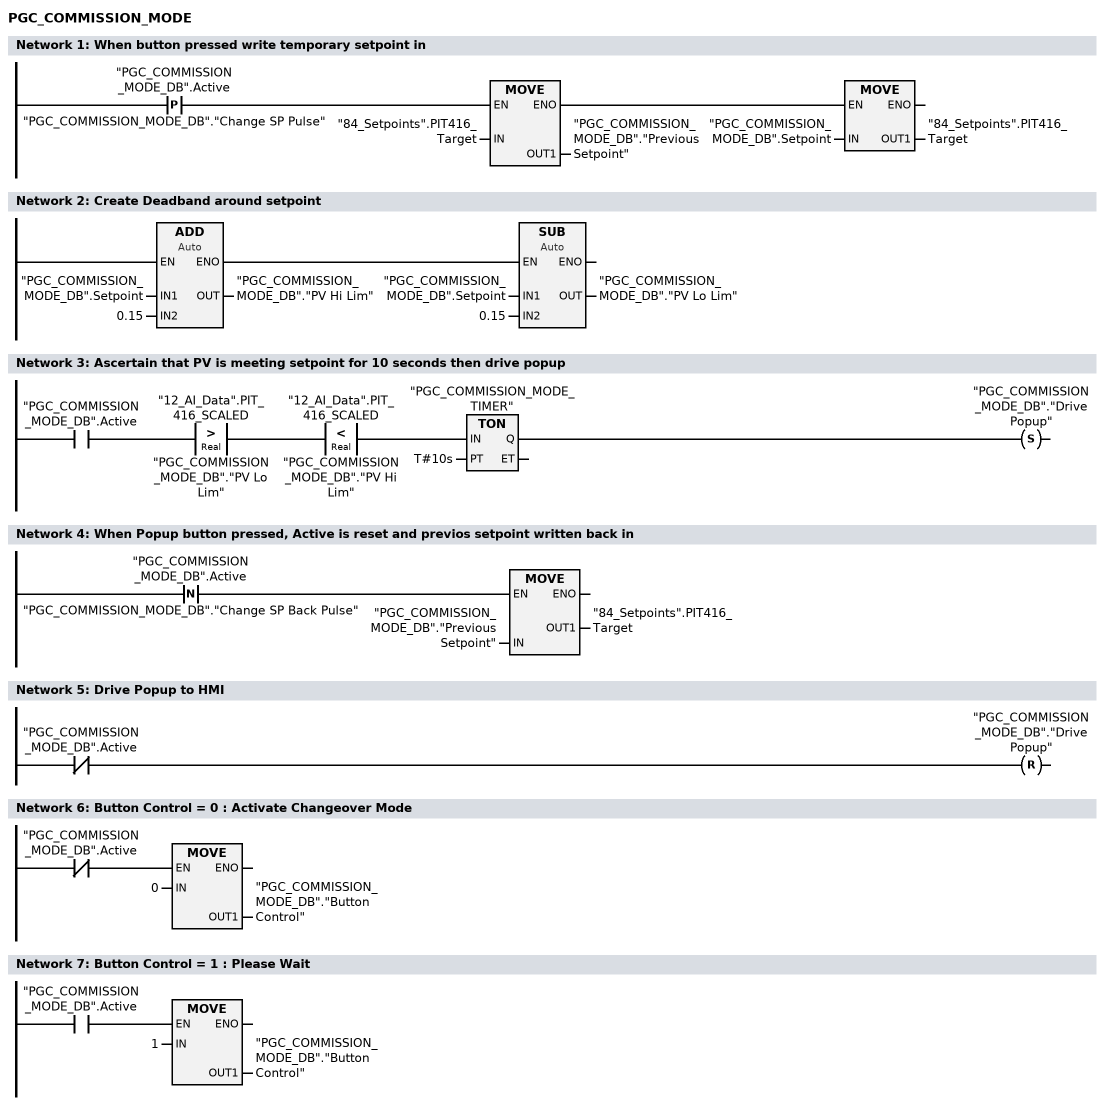
   RUNG wire#powerrail
      P_Contact(operand := "PGC_COMMISSION_MODE_DB".Active, bit := "PGC_COMMISSION_MODE_DB"."Change SP Pulse")
      Move(in := "84_Setpoints".PIT416_Target, out1 => "PGC_COMMISSION_MODE_DB"."Previous Setpoint")
      Move(in := "PGC_COMMISSION_MODE_DB".Setpoint, out1 => "84_Setpoints".PIT416_Target)
   END_RUNG
   // the same network as SCL:
   #_w1 := "PGC_COMMISSION_MODE_DB".Active AND NOT "PGC_COMMISSION_MODE_DB"."Change SP Pulse";   // rising edge of "PGC_COMMISSION_MODE_DB".Active
   "PGC_COMMISSION_MODE_DB"."Change SP Pulse" := "PGC_COMMISSION_MODE_DB".Active;
   IF #_w1 THEN
       "PGC_COMMISSION_MODE_DB"."Previous Setpoint" := "84_Setpoints".PIT416_Target;
       "84_Setpoints".PIT416_Target := "PGC_COMMISSION_MODE_DB".Setpoint;
   END_IF;
END_REGION

REGION Network 2: Create Deadband around setpoint
   RUNG wire#powerrail
      Add(in1 := "PGC_COMMISSION_MODE_DB".Setpoint, in2 := 0.15, out => "PGC_COMMISSION_MODE_DB"."PV Hi Lim")
      Sub(in1 := "PGC_COMMISSION_MODE_DB".Setpoint, in2 := 0.15, out => "PGC_COMMISSION_MODE_DB"."PV Lo Lim")
   END_RUNG
   // the same network as SCL:
   "PGC_COMMISSION_MODE_DB"."PV Hi Lim" := "PGC_COMMISSION_MODE_DB".Setpoint + 0.15;
   "PGC_COMMISSION_MODE_DB"."PV Lo Lim" := "PGC_COMMISSION_MODE_DB".Setpoint - 0.15;
END_REGION

REGION Network 3: Ascertain that PV is meeting setpoint for 10 seconds then drive popup
   "PGC_COMMISSION_MODE_TIMER".TON(IN := "PGC_COMMISSION_MODE_DB".Active AND ("12_AI_Data".PIT_416_SCALED > "PGC_COMMISSION_MODE_DB"."PV Lo Lim") AND ("12_AI_Data".PIT_416_SCALED < "PGC_COMMISSION_MODE_DB"."PV Hi Lim"),
                           PT := T#10s);
   IF "PGC_COMMISSION_MODE_TIMER".Q THEN "PGC_COMMISSION_MODE_DB"."Drive Popup" := TRUE; END_IF;
END_REGION

REGION Network 4: When Popup button pressed, Active is reset and previos setpoint written back in
   RUNG wire#powerrail
      N_Contact(operand := "PGC_COMMISSION_MODE_DB".Active, bit := "PGC_COMMISSION_MODE_DB"."Change SP Back Pulse")
      Move(in := "PGC_COMMISSION_MODE_DB"."Previous Setpoint", out1 => "84_Setpoints".PIT416_Target)
   END_RUNG
   // the same network as SCL:
   #_w1 := NOT "PGC_COMMISSION_MODE_DB".Active AND "PGC_COMMISSION_MODE_DB"."Change SP Back Pulse";   // falling edge of "PGC_COMMISSION_MODE_DB".Active
   "PGC_COMMISSION_MODE_DB"."Change SP Back Pulse" := "PGC_COMMISSION_MODE_DB".Active;
   IF #_w1 THEN "84_Setpoints".PIT416_Target := "PGC_COMMISSION_MODE_DB"."Previous Setpoint"; END_IF;
END_REGION

REGION Network 5: Drive Popup to HMI
   RUNG wire#powerrail
      I_Contact( "PGC_COMMISSION_MODE_DB".Active )
      R_Coil( "PGC_COMMISSION_MODE_DB"."Drive Popup" )
   END_RUNG
   // the same network as SCL:
   IF NOT "PGC_COMMISSION_MODE_DB".Active THEN "PGC_COMMISSION_MODE_DB"."Drive Popup" := FALSE; END_IF;
END_REGION

REGION Network 6: Button Control = 0 : Activate Changeover Mode
   RUNG wire#powerrail
      I_Contact( "PGC_COMMISSION_MODE_DB".Active )
      Move(in := 0, out1 => "PGC_COMMISSION_MODE_DB"."Button Control")
   END_RUNG
   // the same network as SCL:
   IF NOT "PGC_COMMISSION_MODE_DB".Active THEN "PGC_COMMISSION_MODE_DB"."Button Control" := 0; END_IF;
END_REGION

REGION Network 7: Button Control = 1 : Please Wait
   RUNG wire#powerrail
      Contact( "PGC_COMMISSION_MODE_DB".Active )
      Move(in := 1, out1 => "PGC_COMMISSION_MODE_DB"."Button Control")
   END_RUNG
   // the same network as SCL:
   IF "PGC_COMMISSION_MODE_DB".Active THEN "PGC_COMMISSION_MODE_DB"."Button Control" := 1; END_IF;
END_REGION
END_FUNCTION

// folder: 90 - 99 Manual Functions

FUNCTION "90_Manual_Control" : Void   // FC90, LAD
TITLE = Manual Control
{ S7_Optimized_Access := 'TRUE' }
AUTHOR : JHT
VERSION : 0.1
// Code for manual operation of equipment
   VAR_TEMP   // added for the SCL form of the ladder/FBD networks
      _w1 : Bool;
      _w2 : Bool;
      _w3 : Bool;
      _w4 : Bool;
      _w5 : Bool;
      _w6 : Bool;
   END_VAR
BEGIN

REGION Network 1: Q136.0 - Fresh Water Fill Valve Control (CV358)
   // True = Activate, False = NOT
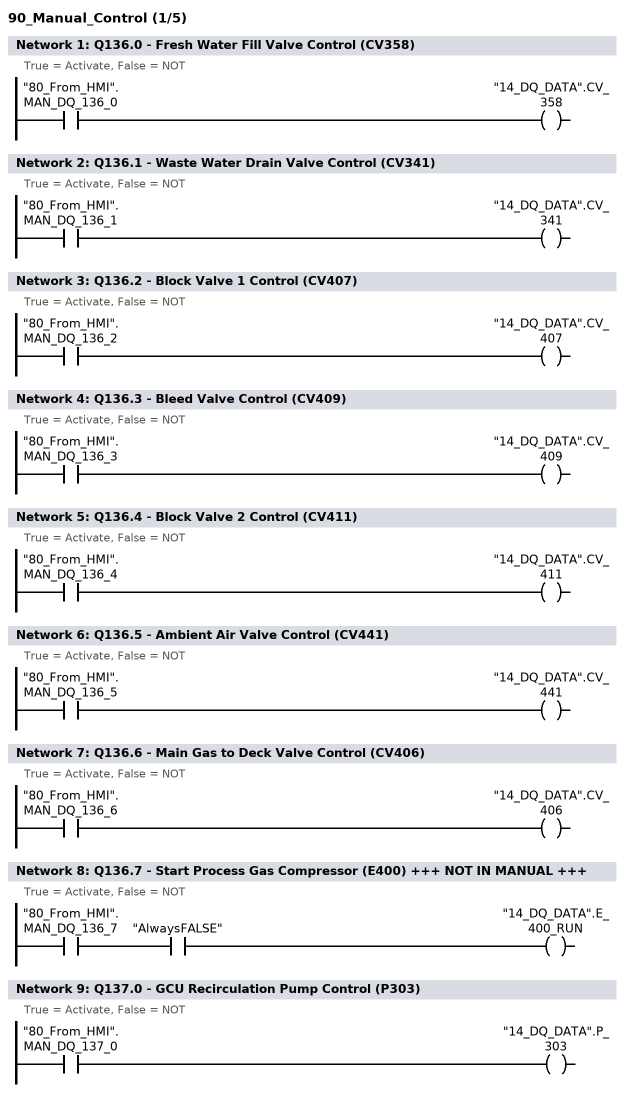
   RUNG wire#powerrail
      Contact( "80_From_HMI".MAN_DQ_136_0 )
      Coil( "14_DQ_DATA".CV_358 )
   END_RUNG
   // the same network as SCL:
   "14_DQ_DATA".CV_358 := "80_From_HMI".MAN_DQ_136_0;
END_REGION

REGION Network 2: Q136.1 - Waste Water Drain Valve Control (CV341)
   // True = Activate, False = NOT
   RUNG wire#powerrail
      Contact( "80_From_HMI".MAN_DQ_136_1 )
      Coil( "14_DQ_DATA".CV_341 )
   END_RUNG
   // the same network as SCL:
   "14_DQ_DATA".CV_341 := "80_From_HMI".MAN_DQ_136_1;
END_REGION

REGION Network 3: Q136.2 - Block Valve 1 Control (CV407)
   // True = Activate, False = NOT
   RUNG wire#powerrail
      Contact( "80_From_HMI".MAN_DQ_136_2 )
      Coil( "14_DQ_DATA".CV_407 )
   END_RUNG
   // the same network as SCL:
   "14_DQ_DATA".CV_407 := "80_From_HMI".MAN_DQ_136_2;
END_REGION

REGION Network 4: Q136.3 - Bleed Valve Control (CV409)
   // True = Activate, False = NOT
   RUNG wire#powerrail
      Contact( "80_From_HMI".MAN_DQ_136_3 )
      Coil( "14_DQ_DATA".CV_409 )
   END_RUNG
   // the same network as SCL:
   "14_DQ_DATA".CV_409 := "80_From_HMI".MAN_DQ_136_3;
END_REGION

REGION Network 5: Q136.4 - Block Valve 2 Control (CV411)
   // True = Activate, False = NOT
   RUNG wire#powerrail
      Contact( "80_From_HMI".MAN_DQ_136_4 )
      Coil( "14_DQ_DATA".CV_411 )
   END_RUNG
   // the same network as SCL:
   "14_DQ_DATA".CV_411 := "80_From_HMI".MAN_DQ_136_4;
END_REGION

REGION Network 6: Q136.5 - Ambient Air Valve Control (CV441)
   // True = Activate, False = NOT
   RUNG wire#powerrail
      Contact( "80_From_HMI".MAN_DQ_136_5 )
      Coil( "14_DQ_DATA".CV_441 )
   END_RUNG
   // the same network as SCL:
   "14_DQ_DATA".CV_441 := "80_From_HMI".MAN_DQ_136_5;
END_REGION

REGION Network 7: Q136.6 - Main Gas to Deck Valve Control (CV406)
   // True = Activate, False = NOT
   RUNG wire#powerrail
      Contact( "80_From_HMI".MAN_DQ_136_6 )
      Coil( "14_DQ_DATA".CV_406 )
   END_RUNG
   // the same network as SCL:
   "14_DQ_DATA".CV_406 := "80_From_HMI".MAN_DQ_136_6;
END_REGION

REGION Network 8: Q136.7 - Start Process Gas Compressor (E400) +++ NOT IN MANUAL +++
   // True = Activate, False = NOT
   RUNG wire#powerrail
      Contact( "80_From_HMI".MAN_DQ_136_7 )
      Contact( "AlwaysFALSE" )
      Coil( "14_DQ_DATA".E_400_RUN )
   END_RUNG
   // the same network as SCL:
   "14_DQ_DATA".E_400_RUN := "80_From_HMI".MAN_DQ_136_7 AND "AlwaysFALSE";
END_REGION

REGION Network 9: Q137.0 - GCU Recirculation Pump Control (P303)
   // True = Activate, False = NOT
   RUNG wire#powerrail
      Contact( "80_From_HMI".MAN_DQ_137_0 )
      Coil( "14_DQ_DATA".P_303 )
   END_RUNG
   // the same network as SCL:
   "14_DQ_DATA".P_303 := "80_From_HMI".MAN_DQ_137_0;
END_REGION

REGION Network 10: Q137.1 - GCU Booster Pump Control (P304)
   // True = Activate, False = NOT
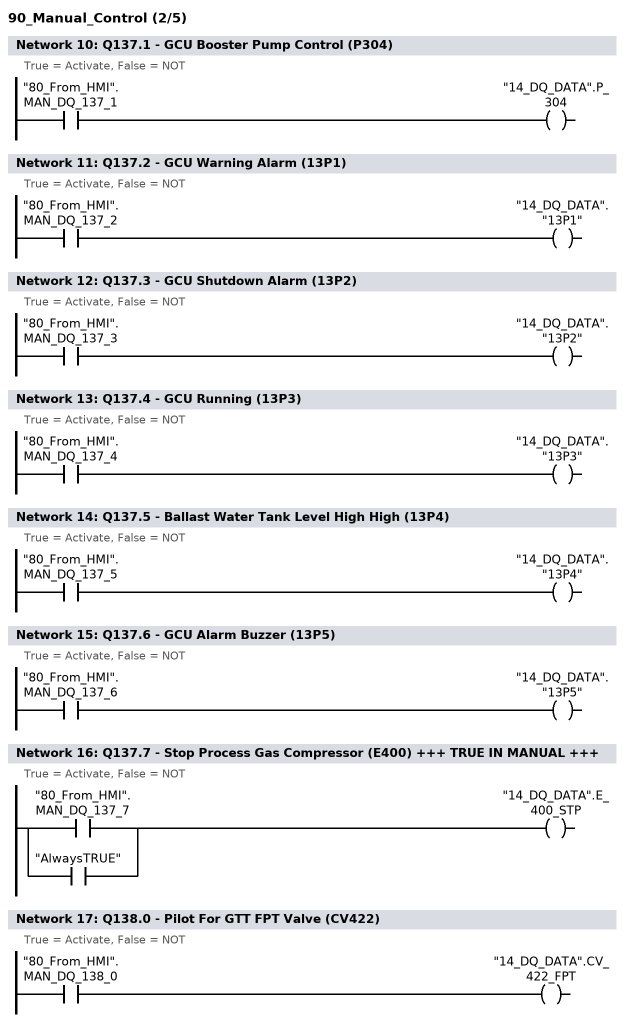
   RUNG wire#powerrail
      Contact( "80_From_HMI".MAN_DQ_137_1 )
      Coil( "14_DQ_DATA".P_304 )
   END_RUNG
   // the same network as SCL:
   "14_DQ_DATA".P_304 := "80_From_HMI".MAN_DQ_137_1;
END_REGION

REGION Network 11: Q137.2 - GCU Warning Alarm (13P1)
   // True = Activate, False = NOT
   RUNG wire#powerrail
      Contact( "80_From_HMI".MAN_DQ_137_2 )
      Coil( "14_DQ_DATA"."13P1" )
   END_RUNG
   // the same network as SCL:
   "14_DQ_DATA"."13P1" := "80_From_HMI".MAN_DQ_137_2;
END_REGION

REGION Network 12: Q137.3 - GCU Shutdown Alarm (13P2)
   // True = Activate, False = NOT
   RUNG wire#powerrail
      Contact( "80_From_HMI".MAN_DQ_137_3 )
      Coil( "14_DQ_DATA"."13P2" )
   END_RUNG
   // the same network as SCL:
   "14_DQ_DATA"."13P2" := "80_From_HMI".MAN_DQ_137_3;
END_REGION

REGION Network 13: Q137.4 - GCU Running (13P3)
   // True = Activate, False = NOT
   RUNG wire#powerrail
      Contact( "80_From_HMI".MAN_DQ_137_4 )
      Coil( "14_DQ_DATA"."13P3" )
   END_RUNG
   // the same network as SCL:
   "14_DQ_DATA"."13P3" := "80_From_HMI".MAN_DQ_137_4;
END_REGION

REGION Network 14: Q137.5 - Ballast Water Tank Level High High (13P4)
   // True = Activate, False = NOT
   RUNG wire#powerrail
      Contact( "80_From_HMI".MAN_DQ_137_5 )
      Coil( "14_DQ_DATA"."13P4" )
   END_RUNG
   // the same network as SCL:
   "14_DQ_DATA"."13P4" := "80_From_HMI".MAN_DQ_137_5;
END_REGION

REGION Network 15: Q137.6 - GCU Alarm Buzzer (13P5)
   // True = Activate, False = NOT
   RUNG wire#powerrail
      Contact( "80_From_HMI".MAN_DQ_137_6 )
      Coil( "14_DQ_DATA"."13P5" )
   END_RUNG
   // the same network as SCL:
   "14_DQ_DATA"."13P5" := "80_From_HMI".MAN_DQ_137_6;
END_REGION

REGION Network 16: Q137.7 - Stop Process Gas Compressor (E400) +++ TRUE IN MANUAL +++
   // True = Activate, False = NOT
   RUNG wire#powerrail
      Contact( "80_From_HMI".MAN_DQ_137_7 )
      wire#w1
      Coil( "14_DQ_DATA".E_400_STP )
   END_RUNG
   RUNG wire#powerrail
      Contact( "AlwaysTRUE" )
   END_RUNG wire#w1
   // the same network as SCL:
   "14_DQ_DATA".E_400_STP := "80_From_HMI".MAN_DQ_137_7 OR "AlwaysTRUE";
END_REGION

REGION Network 17: Q138.0 - Pilot For GTT FPT Valve (CV422)
   // True = Activate, False = NOT
   RUNG wire#powerrail
      Contact( "80_From_HMI".MAN_DQ_138_0 )
      Coil( "14_DQ_DATA".CV_422_FPT )
   END_RUNG
   // the same network as SCL:
   "14_DQ_DATA".CV_422_FPT := "80_From_HMI".MAN_DQ_138_0;
END_REGION

REGION Network 18: Q138.1 - Pilot For GTT 1 Port Valve (CV422)
   // True = Activate, False = NOT
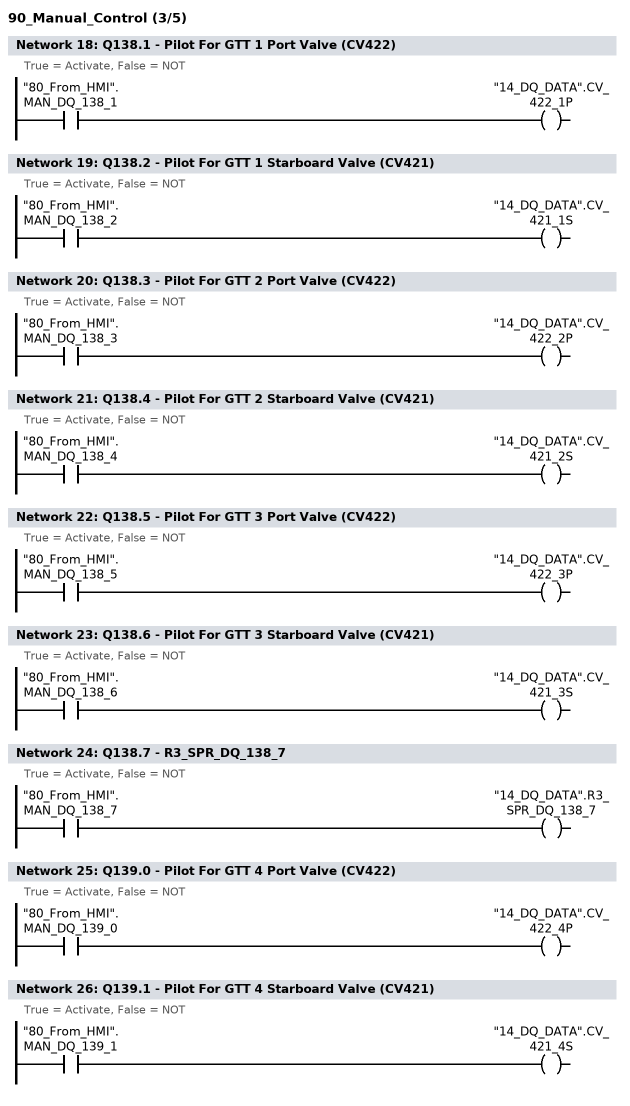
   RUNG wire#powerrail
      Contact( "80_From_HMI".MAN_DQ_138_1 )
      Coil( "14_DQ_DATA".CV_422_1P )
   END_RUNG
   // the same network as SCL:
   "14_DQ_DATA".CV_422_1P := "80_From_HMI".MAN_DQ_138_1;
END_REGION

REGION Network 19: Q138.2 - Pilot For GTT 1 Starboard Valve (CV421)
   // True = Activate, False = NOT
   RUNG wire#powerrail
      Contact( "80_From_HMI".MAN_DQ_138_2 )
      Coil( "14_DQ_DATA".CV_421_1S )
   END_RUNG
   // the same network as SCL:
   "14_DQ_DATA".CV_421_1S := "80_From_HMI".MAN_DQ_138_2;
END_REGION

REGION Network 20: Q138.3 - Pilot For GTT 2 Port Valve (CV422)
   // True = Activate, False = NOT
   RUNG wire#powerrail
      Contact( "80_From_HMI".MAN_DQ_138_3 )
      Coil( "14_DQ_DATA".CV_422_2P )
   END_RUNG
   // the same network as SCL:
   "14_DQ_DATA".CV_422_2P := "80_From_HMI".MAN_DQ_138_3;
END_REGION

REGION Network 21: Q138.4 - Pilot For GTT 2 Starboard Valve (CV421)
   // True = Activate, False = NOT
   RUNG wire#powerrail
      Contact( "80_From_HMI".MAN_DQ_138_4 )
      Coil( "14_DQ_DATA".CV_421_2S )
   END_RUNG
   // the same network as SCL:
   "14_DQ_DATA".CV_421_2S := "80_From_HMI".MAN_DQ_138_4;
END_REGION

REGION Network 22: Q138.5 - Pilot For GTT 3 Port Valve (CV422)
   // True = Activate, False = NOT
   RUNG wire#powerrail
      Contact( "80_From_HMI".MAN_DQ_138_5 )
      Coil( "14_DQ_DATA".CV_422_3P )
   END_RUNG
   // the same network as SCL:
   "14_DQ_DATA".CV_422_3P := "80_From_HMI".MAN_DQ_138_5;
END_REGION

REGION Network 23: Q138.6 - Pilot For GTT 3 Starboard Valve (CV421)
   // True = Activate, False = NOT
   RUNG wire#powerrail
      Contact( "80_From_HMI".MAN_DQ_138_6 )
      Coil( "14_DQ_DATA".CV_421_3S )
   END_RUNG
   // the same network as SCL:
   "14_DQ_DATA".CV_421_3S := "80_From_HMI".MAN_DQ_138_6;
END_REGION

REGION Network 24: Q138.7 - R3_SPR_DQ_138_7
   // True = Activate, False = NOT
   RUNG wire#powerrail
      Contact( "80_From_HMI".MAN_DQ_138_7 )
      Coil( "14_DQ_DATA".R3_SPR_DQ_138_7 )
   END_RUNG
   // the same network as SCL:
   "14_DQ_DATA".R3_SPR_DQ_138_7 := "80_From_HMI".MAN_DQ_138_7;
END_REGION

REGION Network 25: Q139.0 - Pilot For GTT 4 Port Valve (CV422)
   // True = Activate, False = NOT
   RUNG wire#powerrail
      Contact( "80_From_HMI".MAN_DQ_139_0 )
      Coil( "14_DQ_DATA".CV_422_4P )
   END_RUNG
   // the same network as SCL:
   "14_DQ_DATA".CV_422_4P := "80_From_HMI".MAN_DQ_139_0;
END_REGION

REGION Network 26: Q139.1 - Pilot For GTT 4 Starboard Valve (CV421)
   // True = Activate, False = NOT
   RUNG wire#powerrail
      Contact( "80_From_HMI".MAN_DQ_139_1 )
      Coil( "14_DQ_DATA".CV_421_4S )
   END_RUNG
   // the same network as SCL:
   "14_DQ_DATA".CV_421_4S := "80_From_HMI".MAN_DQ_139_1;
END_REGION

REGION Network 27: Q139.2 - Pilot For GTT 5 Port Valve (CV422)
   // True = Activate, False = NOT
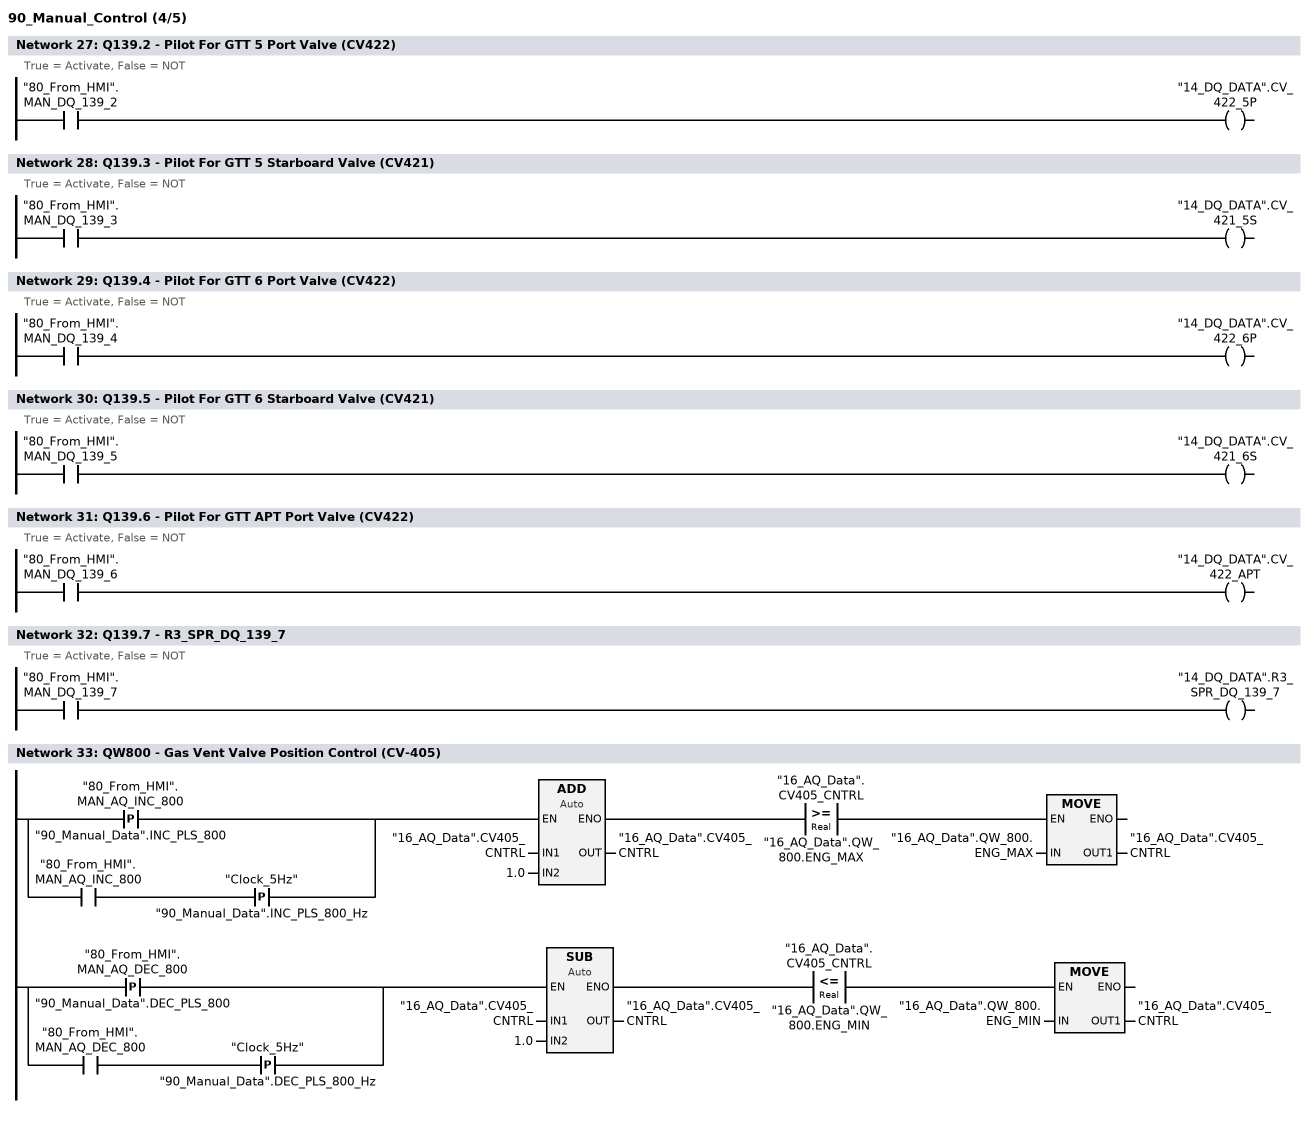
   RUNG wire#powerrail
      Contact( "80_From_HMI".MAN_DQ_139_2 )
      Coil( "14_DQ_DATA".CV_422_5P )
   END_RUNG
   // the same network as SCL:
   "14_DQ_DATA".CV_422_5P := "80_From_HMI".MAN_DQ_139_2;
END_REGION

REGION Network 28: Q139.3 - Pilot For GTT 5 Starboard Valve (CV421)
   // True = Activate, False = NOT
   RUNG wire#powerrail
      Contact( "80_From_HMI".MAN_DQ_139_3 )
      Coil( "14_DQ_DATA".CV_421_5S )
   END_RUNG
   // the same network as SCL:
   "14_DQ_DATA".CV_421_5S := "80_From_HMI".MAN_DQ_139_3;
END_REGION

REGION Network 29: Q139.4 - Pilot For GTT 6 Port Valve (CV422)
   // True = Activate, False = NOT
   RUNG wire#powerrail
      Contact( "80_From_HMI".MAN_DQ_139_4 )
      Coil( "14_DQ_DATA".CV_422_6P )
   END_RUNG
   // the same network as SCL:
   "14_DQ_DATA".CV_422_6P := "80_From_HMI".MAN_DQ_139_4;
END_REGION

REGION Network 30: Q139.5 - Pilot For GTT 6 Starboard Valve (CV421)
   // True = Activate, False = NOT
   RUNG wire#powerrail
      Contact( "80_From_HMI".MAN_DQ_139_5 )
      Coil( "14_DQ_DATA".CV_421_6S )
   END_RUNG
   // the same network as SCL:
   "14_DQ_DATA".CV_421_6S := "80_From_HMI".MAN_DQ_139_5;
END_REGION

REGION Network 31: Q139.6 - Pilot For GTT APT Port Valve (CV422)
   // True = Activate, False = NOT
   RUNG wire#powerrail
      Contact( "80_From_HMI".MAN_DQ_139_6 )
      Coil( "14_DQ_DATA".CV_422_APT )
   END_RUNG
   // the same network as SCL:
   "14_DQ_DATA".CV_422_APT := "80_From_HMI".MAN_DQ_139_6;
END_REGION

REGION Network 32: Q139.7 - R3_SPR_DQ_139_7
   // True = Activate, False = NOT
   RUNG wire#powerrail
      Contact( "80_From_HMI".MAN_DQ_139_7 )
      Coil( "14_DQ_DATA".R3_SPR_DQ_139_7 )
   END_RUNG
   // the same network as SCL:
   "14_DQ_DATA".R3_SPR_DQ_139_7 := "80_From_HMI".MAN_DQ_139_7;
END_REGION

REGION Network 33: QW800 - Gas Vent Valve Position Control (CV-405)
   RUNG wire#powerrail
      P_Contact(operand := "80_From_HMI".MAN_AQ_INC_800, bit := "90_Manual_Data".INC_PLS_800)
      wire#w1
      Add(in1 := "16_AQ_Data".CV405_CNTRL, in2 := 1.0, out => "16_AQ_Data".CV405_CNTRL)
      { S7_Templates := "SrcType := Real" } GE_Contact(in1 := "16_AQ_Data".CV405_CNTRL, in2 := "16_AQ_Data".QW_800.ENG_MAX)
      { S7_GenerateENO := "TRUE" } Move(in := "16_AQ_Data".QW_800.ENG_MAX, out1 => "16_AQ_Data".CV405_CNTRL)
   END_RUNG
   RUNG wire#powerrail
      Contact( "80_From_HMI".MAN_AQ_INC_800 )
      P_Contact(operand := "Clock_5Hz", bit := "90_Manual_Data".INC_PLS_800_Hz)
   END_RUNG wire#w1
   RUNG wire#powerrail
      P_Contact(operand := "80_From_HMI".MAN_AQ_DEC_800, bit := "90_Manual_Data".DEC_PLS_800)
      wire#w2
      Sub(in1 := "16_AQ_Data".CV405_CNTRL, in2 := 1.0, out => "16_AQ_Data".CV405_CNTRL)
      { S7_Templates := "SrcType := Real" } LE_Contact(in1 := "16_AQ_Data".CV405_CNTRL, in2 := "16_AQ_Data".QW_800.ENG_MIN)
      { S7_GenerateENO := "TRUE" } Move(in := "16_AQ_Data".QW_800.ENG_MIN, out1 => "16_AQ_Data".CV405_CNTRL)
   END_RUNG
   RUNG wire#powerrail
      Contact( "80_From_HMI".MAN_AQ_DEC_800 )
      P_Contact(operand := "Clock_5Hz", bit := "90_Manual_Data".DEC_PLS_800_Hz)
   END_RUNG wire#w2
   // the same network as SCL:
   #_w1 := "80_From_HMI".MAN_AQ_INC_800 AND NOT "90_Manual_Data".INC_PLS_800;   // rising edge of "80_From_HMI".MAN_AQ_INC_800
   "90_Manual_Data".INC_PLS_800 := "80_From_HMI".MAN_AQ_INC_800;
   #_w2 := "80_From_HMI".MAN_AQ_INC_800 AND "Clock_5Hz" AND NOT "90_Manual_Data".INC_PLS_800_Hz;   // rising edge of "Clock_5Hz"
   "90_Manual_Data".INC_PLS_800_Hz := "Clock_5Hz";
   #_w3 := #_w1 OR #_w2;
   IF #_w3 THEN "16_AQ_Data".CV405_CNTRL := "16_AQ_Data".CV405_CNTRL + 1.0; END_IF;
   IF #_w3 AND ("16_AQ_Data".CV405_CNTRL >= "16_AQ_Data".QW_800.ENG_MAX) THEN
       "16_AQ_Data".CV405_CNTRL := "16_AQ_Data".QW_800.ENG_MAX;
   END_IF;
   #_w4 := "80_From_HMI".MAN_AQ_DEC_800 AND NOT "90_Manual_Data".DEC_PLS_800;   // rising edge of "80_From_HMI".MAN_AQ_DEC_800
   "90_Manual_Data".DEC_PLS_800 := "80_From_HMI".MAN_AQ_DEC_800;
   #_w5 := "80_From_HMI".MAN_AQ_DEC_800 AND "Clock_5Hz" AND NOT "90_Manual_Data".DEC_PLS_800_Hz;   // rising edge of "Clock_5Hz"
   "90_Manual_Data".DEC_PLS_800_Hz := "Clock_5Hz";
   #_w6 := #_w4 OR #_w5;
   IF #_w6 THEN "16_AQ_Data".CV405_CNTRL := "16_AQ_Data".CV405_CNTRL - 1.0; END_IF;
   IF #_w6 AND ("16_AQ_Data".CV405_CNTRL <= "16_AQ_Data".QW_800.ENG_MIN) THEN
       "16_AQ_Data".CV405_CNTRL := "16_AQ_Data".QW_800.ENG_MIN;
   END_IF;
END_REGION

REGION Network 34: QW802 - Spare Output (Hardware Channel De-activated)
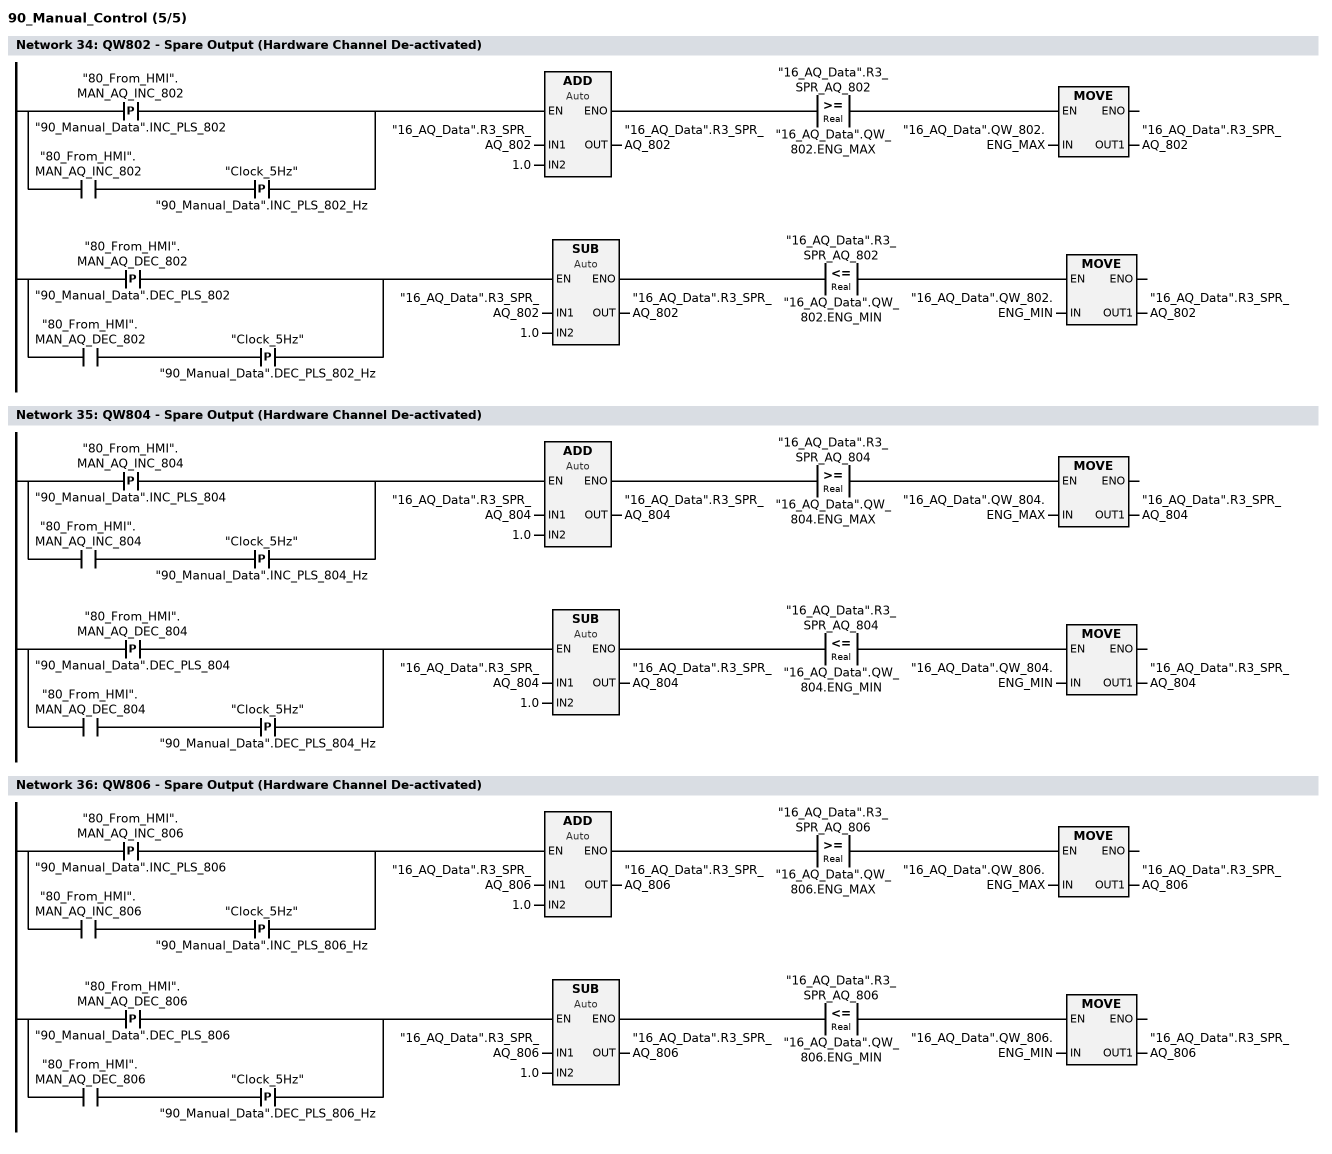
   RUNG wire#powerrail
      P_Contact(operand := "80_From_HMI".MAN_AQ_INC_802, bit := "90_Manual_Data".INC_PLS_802)
      wire#w1
      Add(in1 := "16_AQ_Data".R3_SPR_AQ_802, in2 := 1.0, out => "16_AQ_Data".R3_SPR_AQ_802)
      { S7_Templates := "SrcType := Real" } GE_Contact(in1 := "16_AQ_Data".R3_SPR_AQ_802, in2 := "16_AQ_Data".QW_802.ENG_MAX)
      { S7_GenerateENO := "TRUE" } Move(in := "16_AQ_Data".QW_802.ENG_MAX, out1 => "16_AQ_Data".R3_SPR_AQ_802)
   END_RUNG
   RUNG wire#powerrail
      Contact( "80_From_HMI".MAN_AQ_INC_802 )
      P_Contact(operand := "Clock_5Hz", bit := "90_Manual_Data".INC_PLS_802_Hz)
   END_RUNG wire#w1
   RUNG wire#powerrail
      P_Contact(operand := "80_From_HMI".MAN_AQ_DEC_802, bit := "90_Manual_Data".DEC_PLS_802)
      wire#w2
      Sub(in1 := "16_AQ_Data".R3_SPR_AQ_802, in2 := 1.0, out => "16_AQ_Data".R3_SPR_AQ_802)
      { S7_Templates := "SrcType := Real" } LE_Contact(in1 := "16_AQ_Data".R3_SPR_AQ_802, in2 := "16_AQ_Data".QW_802.ENG_MIN)
      { S7_GenerateENO := "TRUE" } Move(in := "16_AQ_Data".QW_802.ENG_MIN, out1 => "16_AQ_Data".R3_SPR_AQ_802)
   END_RUNG
   RUNG wire#powerrail
      Contact( "80_From_HMI".MAN_AQ_DEC_802 )
      P_Contact(operand := "Clock_5Hz", bit := "90_Manual_Data".DEC_PLS_802_Hz)
   END_RUNG wire#w2
   // the same network as SCL:
   #_w1 := "80_From_HMI".MAN_AQ_INC_802 AND NOT "90_Manual_Data".INC_PLS_802;   // rising edge of "80_From_HMI".MAN_AQ_INC_802
   "90_Manual_Data".INC_PLS_802 := "80_From_HMI".MAN_AQ_INC_802;
   #_w2 := "80_From_HMI".MAN_AQ_INC_802 AND "Clock_5Hz" AND NOT "90_Manual_Data".INC_PLS_802_Hz;   // rising edge of "Clock_5Hz"
   "90_Manual_Data".INC_PLS_802_Hz := "Clock_5Hz";
   #_w3 := #_w1 OR #_w2;
   IF #_w3 THEN "16_AQ_Data".R3_SPR_AQ_802 := "16_AQ_Data".R3_SPR_AQ_802 + 1.0; END_IF;
   IF #_w3 AND ("16_AQ_Data".R3_SPR_AQ_802 >= "16_AQ_Data".QW_802.ENG_MAX) THEN
       "16_AQ_Data".R3_SPR_AQ_802 := "16_AQ_Data".QW_802.ENG_MAX;
   END_IF;
   #_w4 := "80_From_HMI".MAN_AQ_DEC_802 AND NOT "90_Manual_Data".DEC_PLS_802;   // rising edge of "80_From_HMI".MAN_AQ_DEC_802
   "90_Manual_Data".DEC_PLS_802 := "80_From_HMI".MAN_AQ_DEC_802;
   #_w5 := "80_From_HMI".MAN_AQ_DEC_802 AND "Clock_5Hz" AND NOT "90_Manual_Data".DEC_PLS_802_Hz;   // rising edge of "Clock_5Hz"
   "90_Manual_Data".DEC_PLS_802_Hz := "Clock_5Hz";
   #_w6 := #_w4 OR #_w5;
   IF #_w6 THEN "16_AQ_Data".R3_SPR_AQ_802 := "16_AQ_Data".R3_SPR_AQ_802 - 1.0; END_IF;
   IF #_w6 AND ("16_AQ_Data".R3_SPR_AQ_802 <= "16_AQ_Data".QW_802.ENG_MIN) THEN
       "16_AQ_Data".R3_SPR_AQ_802 := "16_AQ_Data".QW_802.ENG_MIN;
   END_IF;
END_REGION

REGION Network 35: QW804 - Spare Output (Hardware Channel De-activated)
   RUNG wire#powerrail
      P_Contact(operand := "80_From_HMI".MAN_AQ_INC_804, bit := "90_Manual_Data".INC_PLS_804)
      wire#w1
      Add(in1 := "16_AQ_Data".R3_SPR_AQ_804, in2 := 1.0, out => "16_AQ_Data".R3_SPR_AQ_804)
      { S7_Templates := "SrcType := Real" } GE_Contact(in1 := "16_AQ_Data".R3_SPR_AQ_804, in2 := "16_AQ_Data".QW_804.ENG_MAX)
      { S7_GenerateENO := "TRUE" } Move(in := "16_AQ_Data".QW_804.ENG_MAX, out1 => "16_AQ_Data".R3_SPR_AQ_804)
   END_RUNG
   RUNG wire#powerrail
      Contact( "80_From_HMI".MAN_AQ_INC_804 )
      P_Contact(operand := "Clock_5Hz", bit := "90_Manual_Data".INC_PLS_804_Hz)
   END_RUNG wire#w1
   RUNG wire#powerrail
      P_Contact(operand := "80_From_HMI".MAN_AQ_DEC_804, bit := "90_Manual_Data".DEC_PLS_804)
      wire#w2
      Sub(in1 := "16_AQ_Data".R3_SPR_AQ_804, in2 := 1.0, out => "16_AQ_Data".R3_SPR_AQ_804)
      { S7_Templates := "SrcType := Real" } LE_Contact(in1 := "16_AQ_Data".R3_SPR_AQ_804, in2 := "16_AQ_Data".QW_804.ENG_MIN)
      { S7_GenerateENO := "TRUE" } Move(in := "16_AQ_Data".QW_804.ENG_MIN, out1 => "16_AQ_Data".R3_SPR_AQ_804)
   END_RUNG
   RUNG wire#powerrail
      Contact( "80_From_HMI".MAN_AQ_DEC_804 )
      P_Contact(operand := "Clock_5Hz", bit := "90_Manual_Data".DEC_PLS_804_Hz)
   END_RUNG wire#w2
   // the same network as SCL:
   #_w1 := "80_From_HMI".MAN_AQ_INC_804 AND NOT "90_Manual_Data".INC_PLS_804;   // rising edge of "80_From_HMI".MAN_AQ_INC_804
   "90_Manual_Data".INC_PLS_804 := "80_From_HMI".MAN_AQ_INC_804;
   #_w2 := "80_From_HMI".MAN_AQ_INC_804 AND "Clock_5Hz" AND NOT "90_Manual_Data".INC_PLS_804_Hz;   // rising edge of "Clock_5Hz"
   "90_Manual_Data".INC_PLS_804_Hz := "Clock_5Hz";
   #_w3 := #_w1 OR #_w2;
   IF #_w3 THEN "16_AQ_Data".R3_SPR_AQ_804 := "16_AQ_Data".R3_SPR_AQ_804 + 1.0; END_IF;
   IF #_w3 AND ("16_AQ_Data".R3_SPR_AQ_804 >= "16_AQ_Data".QW_804.ENG_MAX) THEN
       "16_AQ_Data".R3_SPR_AQ_804 := "16_AQ_Data".QW_804.ENG_MAX;
   END_IF;
   #_w4 := "80_From_HMI".MAN_AQ_DEC_804 AND NOT "90_Manual_Data".DEC_PLS_804;   // rising edge of "80_From_HMI".MAN_AQ_DEC_804
   "90_Manual_Data".DEC_PLS_804 := "80_From_HMI".MAN_AQ_DEC_804;
   #_w5 := "80_From_HMI".MAN_AQ_DEC_804 AND "Clock_5Hz" AND NOT "90_Manual_Data".DEC_PLS_804_Hz;   // rising edge of "Clock_5Hz"
   "90_Manual_Data".DEC_PLS_804_Hz := "Clock_5Hz";
   #_w6 := #_w4 OR #_w5;
   IF #_w6 THEN "16_AQ_Data".R3_SPR_AQ_804 := "16_AQ_Data".R3_SPR_AQ_804 - 1.0; END_IF;
   IF #_w6 AND ("16_AQ_Data".R3_SPR_AQ_804 <= "16_AQ_Data".QW_804.ENG_MIN) THEN
       "16_AQ_Data".R3_SPR_AQ_804 := "16_AQ_Data".QW_804.ENG_MIN;
   END_IF;
END_REGION

REGION Network 36: QW806 - Spare Output (Hardware Channel De-activated)
   RUNG wire#powerrail
      P_Contact(operand := "80_From_HMI".MAN_AQ_INC_806, bit := "90_Manual_Data".INC_PLS_806)
      wire#w1
      Add(in1 := "16_AQ_Data".R3_SPR_AQ_806, in2 := 1.0, out => "16_AQ_Data".R3_SPR_AQ_806)
      { S7_Templates := "SrcType := Real" } GE_Contact(in1 := "16_AQ_Data".R3_SPR_AQ_806, in2 := "16_AQ_Data".QW_806.ENG_MAX)
      { S7_GenerateENO := "TRUE" } Move(in := "16_AQ_Data".QW_806.ENG_MAX, out1 => "16_AQ_Data".R3_SPR_AQ_806)
   END_RUNG
   RUNG wire#powerrail
      Contact( "80_From_HMI".MAN_AQ_INC_806 )
      P_Contact(operand := "Clock_5Hz", bit := "90_Manual_Data".INC_PLS_806_Hz)
   END_RUNG wire#w1
   RUNG wire#powerrail
      P_Contact(operand := "80_From_HMI".MAN_AQ_DEC_806, bit := "90_Manual_Data".DEC_PLS_806)
      wire#w2
      Sub(in1 := "16_AQ_Data".R3_SPR_AQ_806, in2 := 1.0, out => "16_AQ_Data".R3_SPR_AQ_806)
      { S7_Templates := "SrcType := Real" } LE_Contact(in1 := "16_AQ_Data".R3_SPR_AQ_806, in2 := "16_AQ_Data".QW_806.ENG_MIN)
      { S7_GenerateENO := "TRUE" } Move(in := "16_AQ_Data".QW_806.ENG_MIN, out1 => "16_AQ_Data".R3_SPR_AQ_806)
   END_RUNG
   RUNG wire#powerrail
      Contact( "80_From_HMI".MAN_AQ_DEC_806 )
      P_Contact(operand := "Clock_5Hz", bit := "90_Manual_Data".DEC_PLS_806_Hz)
   END_RUNG wire#w2
   // the same network as SCL:
   #_w1 := "80_From_HMI".MAN_AQ_INC_806 AND NOT "90_Manual_Data".INC_PLS_806;   // rising edge of "80_From_HMI".MAN_AQ_INC_806
   "90_Manual_Data".INC_PLS_806 := "80_From_HMI".MAN_AQ_INC_806;
   #_w2 := "80_From_HMI".MAN_AQ_INC_806 AND "Clock_5Hz" AND NOT "90_Manual_Data".INC_PLS_806_Hz;   // rising edge of "Clock_5Hz"
   "90_Manual_Data".INC_PLS_806_Hz := "Clock_5Hz";
   #_w3 := #_w1 OR #_w2;
   IF #_w3 THEN "16_AQ_Data".R3_SPR_AQ_806 := "16_AQ_Data".R3_SPR_AQ_806 + 1.0; END_IF;
   IF #_w3 AND ("16_AQ_Data".R3_SPR_AQ_806 >= "16_AQ_Data".QW_806.ENG_MAX) THEN
       "16_AQ_Data".R3_SPR_AQ_806 := "16_AQ_Data".QW_806.ENG_MAX;
   END_IF;
   #_w4 := "80_From_HMI".MAN_AQ_DEC_806 AND NOT "90_Manual_Data".DEC_PLS_806;   // rising edge of "80_From_HMI".MAN_AQ_DEC_806
   "90_Manual_Data".DEC_PLS_806 := "80_From_HMI".MAN_AQ_DEC_806;
   #_w5 := "80_From_HMI".MAN_AQ_DEC_806 AND "Clock_5Hz" AND NOT "90_Manual_Data".DEC_PLS_806_Hz;   // rising edge of "Clock_5Hz"
   "90_Manual_Data".DEC_PLS_806_Hz := "Clock_5Hz";
   #_w6 := #_w4 OR #_w5;
   IF #_w6 THEN "16_AQ_Data".R3_SPR_AQ_806 := "16_AQ_Data".R3_SPR_AQ_806 - 1.0; END_IF;
   IF #_w6 AND ("16_AQ_Data".R3_SPR_AQ_806 <= "16_AQ_Data".QW_806.ENG_MIN) THEN
       "16_AQ_Data".R3_SPR_AQ_806 := "16_AQ_Data".QW_806.ENG_MIN;
   END_IF;
END_REGION
END_FUNCTION

(* ===== HMI "HMI_RT_1" =====
system functions are stored by id; their names below are inferred from use
connection "IGG PLC Comms": ETHERNET, S7_1500_OMS
connection "BC PLC Comms": ETHERNET, S7_1500_OMS
connection "BWTS PLC Comms": ETHERNET, S7_1500_OMS

